HMI tags "PackTags"
   "PackTags.Admin.ProdProcessedCount[0].Count" : DInt = PLC PackTags.Admin.ProdProcessedCount[0].Count, 1 s   // Total Number of Products Through Machine / Número total de productos a través de la máquina
   "PackTags.Admin.ProdDefectiveCount[0].Count" : DInt = PLC PackTags.Admin.ProdDefectiveCount[0].Count, 1 s   // Total Number of Defective Products the Machine Processed (Reject Total ) / Número total de productos defectuosos procesados por la máquina (rechazo total)
   "PackTags.Admin.StopReason.ID" : DInt = PLC PackTags.Admin.StopReason.ID, 1 s   // Unique value assigned to each alarm
   "PackTags.Admin.StopReason.Value" : DInt = PLC PackTags.Admin.StopReason.Value, 1 s   // The Alarm Message number is a value that is associated to the alarm allowing for user specific detail or to break down the Alarm.ID to greater detail
   "PackTags.Admin.ProdProcessedCount[0].Unit" : String[5] = PLC PackTags.Admin.ProdProcessedCount[0].Unit, 1 s
   "PackTags.Admin.StatesDisabled" : DInt = PLC PackTags.Admin.StatesDisabled, 1 s
   "PackTags.Command.CmdChangeRequest" : Bool = PLC PackTags.Command.CmdChangeRequest, 1 s
   "PackTags.Command.CntrlCmd" : DInt = PLC PackTags.Command.CntrlCmd, 1 s
   "PackTags.Command.MachSpeed" : Real = PLC PackTags.Command.MachSpeed AT %DB1.DBD0, 1 s
   "PackTags.Command.UnitMode" : DInt = PLC PackTags.Command.UnitMode, 1 s
   "PackTags.Command.UnitModeChangeRequest" : Bool = PLC PackTags.Command.UnitModeChangeRequest, 1 s
   "PackML.remoteCommandEnable" : Bool = PLC PackML.remoteCommandEnable, 1 s
   "PackTags.Status.CurMachSpeed" : Real = PLC PackTags.Status.CurMachSpeed, 1 s
   "PackTags.Status.EquipmentInterlock.Blocked" : Bool = PLC PackTags.Status.EquipmentInterlock.Blocked, 1 s
   "PackTags.Status.EquipmentInterlock.Starved" : Bool = PLC PackTags.Status.EquipmentInterlock.Starved, 1 s
   "PackTags.Status.MachSpeed" : Real = PLC PackTags.Status.MachSpeed, 1 s
   "PackTags.Status.StateCurrent" : DInt = PLC PackTags.Status.StateCurrent, 500 ms
   "PackTags.Status.StateCurrentName" : String[16] = PLC PackTags.Status.StateCurrentName, 1 s
   "PackTags.Status.UnitModeCurrent" : DInt = PLC PackTags.Status.UnitModeCurrent, 1 s
   "PackTags.Status.UnitModeCurrentName" : String[18] = PLC PackTags.Status.UnitModeCurrentName, 1 s
   "PackML.Cmd.Mode.Maintenance" : Bool = PLC PackML.Cmd.Mode.Maintenance AT %DB1.DBX0.0, 1 s
   "PackML.Cmd.Mode.Manual" : Bool = PLC PackML.Cmd.Mode.Manual, 1 s
   "PackML.Cmd.Mode.Production" : Bool = PLC PackML.Cmd.Mode.Production, 1 s
   "PackML.Cmd.Mode.UserMode01" : Bool = PLC PackML.Cmd.Mode.UserMode01 AT %DB1.DBX0.0, 1 s
   "PackTags.Admin.AlarmExtent" : DInt = PLC PackTags.Admin.AlarmExtent, 1 s
   "PackTags.Admin.MachDesignSpeed" : Real = PLC PackTags.Admin.MachDesignSpeed AT %DB1.DBX0.0, 1 s
   "PackTags.Admin.ProdConsumedCount[0].AccCount" : DInt = PLC PackTags.Admin.ProdConsumedCount[0].AccCount, 1 s
   "PackTags.Admin.ProdConsumedCount[0].Count" : DInt = PLC PackTags.Admin.ProdConsumedCount[0].Count, 1 s
   "PackTags.Admin.ProdConsumedCount[0].Name" : String[24] = PLC PackTags.Admin.ProdConsumedCount[0].Name, 1 s
   "PackTags.Admin.ProdConsumedCount[0].Unit" : String[5] = PLC PackTags.Admin.ProdConsumedCount[0].Unit, 1 s
   "PackTags.Admin.ProdDefectiveCount[0].AccCount" : DInt = PLC PackTags.Admin.ProdDefectiveCount[0].AccCount, 1 s
   "PackTags.Admin.ProdDefectiveCount[0].Name" : String[24] = PLC PackTags.Admin.ProdDefectiveCount[0].Name, 1 s
   "PackTags.Admin.ProdDefectiveCount[0].Unit" : String[5] = PLC PackTags.Admin.ProdDefectiveCount[0].Unit, 1 s
   "PackTags.Admin.ProdProcessedCount[0].AccCount" : DInt = PLC PackTags.Admin.ProdProcessedCount[0].AccCount, 1 s
   "PackTags.Admin.ProdProcessedCount[0].Name" : String[24] = PLC PackTags.Admin.ProdProcessedCount[0].Name, 1 s
   "PackTags.Status.MaterialInterlock" : DWord = PLC PackTags.Status.MaterialInterlock AT %DB1.DBD0, 1 s

HMI tags "Tag table_PackTags_Times"
   "HMI_Data.resetPackMLTimers" : Bool = PLC HMI_Data.resetPackMLTimers, 500 ms   // Reset the PackML Timer values when set (1). / Restablezca los valores del temporizador PackML cuando se establece (1).
   "HMI_Data.modeCumulativeTime" : DInt = PLC HMI_Data.modeCumulativeTime, 1 s
   "HMI_Data.State_Current_Times[1]" : DInt = PLC HMI_Data.State_Current_Times[1], 1 s
   "HMI_Data.State_Current_Times[2]" : DInt = PLC HMI_Data.State_Current_Times[2], 1 s
   "HMI_Data.State_Current_Times[3]" : DInt = PLC HMI_Data.State_Current_Times[3], 1 s
   "HMI_Data.State_Current_Times[4]" : DInt = PLC HMI_Data.State_Current_Times[4], 1 s
   "HMI_Data.State_Current_Times[5]" : DInt = PLC HMI_Data.State_Current_Times[5], 1 s
   "HMI_Data.State_Current_Times[6]" : DInt = PLC HMI_Data.State_Current_Times[6], 1 s
   "HMI_Data.State_Current_Times[7]" : DInt = PLC HMI_Data.State_Current_Times[7], 1 s
   "HMI_Data.State_Current_Times[8]" : DInt = PLC HMI_Data.State_Current_Times[8], 1 s
   "HMI_Data.State_Current_Times[9]" : DInt = PLC HMI_Data.State_Current_Times[9], 1 s
   "HMI_Data.State_Current_Times[10]" : DInt = PLC HMI_Data.State_Current_Times[10], 1 s
   "HMI_Data.State_Current_Times[11]" : DInt = PLC HMI_Data.State_Current_Times[11], 1 s
   "HMI_Data.State_Current_Times[12]" : DInt = PLC HMI_Data.State_Current_Times[12], 1 s
   "HMI_Data.State_Current_Times[13]" : DInt = PLC HMI_Data.State_Current_Times[13], 1 s
   "HMI_Data.State_Current_Times[14]" : DInt = PLC HMI_Data.State_Current_Times[14], 1 s
   "HMI_Data.State_Current_Times[15]" : DInt = PLC HMI_Data.State_Current_Times[15], 1 s
   "HMI_Data.State_Current_Times[16]" : DInt = PLC HMI_Data.State_Current_Times[16], 1 s
   "HMI_Data.State_Current_Times[17]" : DInt = PLC HMI_Data.State_Current_Times[17], 1 s
   "HMI_Data.State_Cumulative_Times[1]" : DInt = PLC HMI_Data.State_Cumulative_Times[1], 1 s
   "HMI_Data.State_Cumulative_Times[2]" : DInt = PLC HMI_Data.State_Cumulative_Times[2], 1 s
   "HMI_Data.State_Cumulative_Times[3]" : DInt = PLC HMI_Data.State_Cumulative_Times[3], 1 s
   "HMI_Data.State_Cumulative_Times[4]" : DInt = PLC HMI_Data.State_Cumulative_Times[4], 1 s
   "HMI_Data.State_Cumulative_Times[5]" : DInt = PLC HMI_Data.State_Cumulative_Times[5], 1 s
   "HMI_Data.State_Cumulative_Times[6]" : DInt = PLC HMI_Data.State_Cumulative_Times[6], 1 s
   "HMI_Data.State_Cumulative_Times[7]" : DInt = PLC HMI_Data.State_Cumulative_Times[7], 1 s
   "HMI_Data.State_Cumulative_Times[8]" : DInt = PLC HMI_Data.State_Cumulative_Times[8], 1 s
   "HMI_Data.State_Cumulative_Times[9]" : DInt = PLC HMI_Data.State_Cumulative_Times[9], 1 s
   "HMI_Data.State_Cumulative_Times[10]" : DInt = PLC HMI_Data.State_Cumulative_Times[10], 1 s
   "HMI_Data.State_Cumulative_Times[11]" : DInt = PLC HMI_Data.State_Cumulative_Times[11], 1 s
   "HMI_Data.State_Cumulative_Times[12]" : DInt = PLC HMI_Data.State_Cumulative_Times[12], 1 s
   "HMI_Data.State_Cumulative_Times[13]" : DInt = PLC HMI_Data.State_Cumulative_Times[13], 1 s
   "HMI_Data.State_Cumulative_Times[14]" : DInt = PLC HMI_Data.State_Cumulative_Times[14], 1 s
   "HMI_Data.State_Cumulative_Times[15]" : DInt = PLC HMI_Data.State_Cumulative_Times[15], 1 s
   "HMI_Data.State_Cumulative_Times[16]" : DInt = PLC HMI_Data.State_Cumulative_Times[16], 1 s
   "HMI_Data.State_Cumulative_Times[17]" : DInt = PLC HMI_Data.State_Cumulative_Times[17], 1 s
   "PackTags.Admin.ModeCurrentTime[1]" : DInt = PLC PackTags.Admin.ModeCurrentTime[1], 1 s
   "PackTags.Admin.ModeCurrentTime[2]" : DInt = PLC PackTags.Admin.ModeCurrentTime[2], 1 s
   "PackTags.Admin.ModeCurrentTime[3]" : DInt = PLC PackTags.Admin.ModeCurrentTime[3], 1 s
   "PackTags.Admin.ModeCurrentTime[4]" : DInt = PLC PackTags.Admin.ModeCurrentTime[4], 1 s
   "PackTags.Admin.ModeCumulativeTime[1]" : DInt = PLC PackTags.Admin.ModeCumulativeTime[1], 1 s
   "PackTags.Admin.ModeCumulativeTime[2]" : DInt = PLC PackTags.Admin.ModeCumulativeTime[2], 1 s
   "PackTags.Admin.ModeCumulativeTime[3]" : DInt = PLC PackTags.Admin.ModeCumulativeTime[3], 1 s
   "PackTags.Admin.ModeCumulativeTime[4]" : DInt = PLC PackTags.Admin.ModeCumulativeTime[4], 1 s
   "PackTags.Admin.AccTimeSinceLastReset" : DInt = PLC PackTags.Admin.AccTimeSinceLastReset, 1 s

HMI tags "Tag table_Event_Warning_SortFilter"
   "HMI_Data.EMSortDisableWarning.EM00" : Bool = PLC HMI_Data.EMSortDisableWarning.EM00, 1 s   // If bool is reset, then EMxx sort filter is enabled, else it's disabled. / If bool is reset, then EMxx is sort filter is enabled, else it's disabled.
   "HMI_Data.EMSortDisableWarning.EM01" : Bool = PLC HMI_Data.EMSortDisableWarning.EM01, 1 s   // If bool is reset, then EMxx sort filter is enabled, else it's disabled. / If bool is reset, then EMxx is sort filter is enabled, else it's disabled.
   "HMI_Data.EMSortDisableWarning.EM02" : Bool = PLC HMI_Data.EMSortDisableWarning.EM02, 1 s   // If bool is reset, then EMxx sort filter is enabled, else it's disabled. / If bool is reset, then EMxx is sort filter is enabled, else it's disabled.
   "HMI_Data.EMSortDisableWarning.EM03" : Bool = PLC HMI_Data.EMSortDisableWarning.EM03, 1 s   // If bool is reset, then EMxx sort filter is enabled, else it's disabled. / If bool is reset, then EMxx is sort filter is enabled, else it's disabled.
   "HMI_Data.EMSortDisableWarning.EM04" : Bool = PLC HMI_Data.EMSortDisableWarning.EM04, 1 s   // If bool is reset, then EMxx sort filter is enabled, else it's disabled. / If bool is reset, then EMxx is sort filter is enabled, else it's disabled.
   "HMI_Data.EMSortDisableWarning.EM05" : Bool = PLC HMI_Data.EMSortDisableWarning.EM05, 1 s   // If bool is reset, then EMxx sort filter is enabled, else it's disabled. / If bool is reset, then EMxx is sort filter is enabled, else it's disabled.
   "HMI_Data.EMSortDisableWarning.EM06" : Bool = PLC HMI_Data.EMSortDisableWarning.EM06, 1 s   // If bool is reset, then EMxx sort filter is enabled, else it's disabled. / If bool is reset, then EMxx is sort filter is enabled, else it's disabled.
   "HMI_Data.EMSortDisableWarning.EM07" : Bool = PLC HMI_Data.EMSortDisableWarning.EM07, 1 s   // If bool is reset, then EMxx sort filter is enabled, else it's disabled. / If bool is reset, then EMxx is sort filter is enabled, else it's disabled.
   "HMI_Data.EMSortDisableWarning.EM08" : Bool = PLC HMI_Data.EMSortDisableWarning.EM08, 1 s   // If bool is reset, then EMxx sort filter is enabled, else it's disabled. / If bool is reset, then EMxx is sort filter is enabled, else it's disabled.
   "HMI_Data.EMSortDisableWarning.EM09" : Bool = PLC HMI_Data.EMSortDisableWarning.EM09, 1 s   // If bool is reset, then EMxx sort filter is enabled, else it's disabled. / If bool is reset, then EMxx is sort filter is enabled, else it's disabled.
   "HMI_Data.EMSortDisableWarning.EM10" : Bool = PLC HMI_Data.EMSortDisableWarning.EM10, 1 s   // If bool is reset, then EMxx sort filter is enabled, else it's disabled. / If bool is reset, then EMxx is sort filter is enabled, else it's disabled.
   "HMI_Data.EMSortDisableWarning.Unit" : Bool = PLC HMI_Data.EMSortDisableWarning.Unit, 1 s   // If bool is reset, then Unit sort filter is enabled, else it's disabled. / If bool is reset, then EMxx is sort filter is enabled, else it's disabled.

HMI tags "Tag table_Event_Warning"
   "HMI_Data.warningSortedList[0]" : CPG_typeEvent = PLC HMI_Data.warningSortedList[0], 1 s
   "HMI_Data.warningSortedList[1]" : CPG_typeEvent = PLC HMI_Data.warningSortedList[1], 1 s
   "HMI_Data.warningSortedList[2]" : CPG_typeEvent = PLC HMI_Data.warningSortedList[2], 1 s
   "HMI_Data.warningSortedList[3]" : CPG_typeEvent = PLC HMI_Data.warningSortedList[3], 1 s
   "HMI_Data.warningSortedList[4]" : CPG_typeEvent = PLC HMI_Data.warningSortedList[4], 1 s
   "HMI_Data.warningSortedList[5]" : CPG_typeEvent = PLC HMI_Data.warningSortedList[5], 1 s
   "HMI_Data.warningSortedList[6]" : CPG_typeEvent = PLC HMI_Data.warningSortedList[6], 1 s
   "HMI_Data.warningSortedList[7]" : CPG_typeEvent = PLC HMI_Data.warningSortedList[7], 1 s
   "HMI_Data.warningSortedList[8]" : CPG_typeEvent = PLC HMI_Data.warningSortedList[8], 1 s
   "HMI_Data.warningSortedList[9]" : CPG_typeEvent = PLC HMI_Data.warningSortedList[9], 1 s
   "HMI_Data.warningSortedList[10]" : CPG_typeEvent = PLC HMI_Data.warningSortedList[10], 1 s
   "HMI_Data.warningSortedList[11]" : CPG_typeEvent = PLC HMI_Data.warningSortedList[11], 1 s
   "HMI_Data.warningSortedList[12]" : CPG_typeEvent = PLC HMI_Data.warningSortedList[12], 1 s
   "HMI_Data.warningSortedList[13]" : CPG_typeEvent = PLC HMI_Data.warningSortedList[13], 1 s
   "HMI_Data.warningSortedList[14]" : CPG_typeEvent = PLC HMI_Data.warningSortedList[14], 1 s
   "HMI_Data.warningSortedList[15]" : CPG_typeEvent = PLC HMI_Data.warningSortedList[15], 1 s
   "HMI_Data.warningSortedList[16]" : CPG_typeEvent = PLC HMI_Data.warningSortedList[16], 1 s
   "HMI_Data.warningSortedList[17]" : CPG_typeEvent = PLC HMI_Data.warningSortedList[17], 1 s
   "HMI_Data.warningSortedList[18]" : CPG_typeEvent = PLC HMI_Data.warningSortedList[18], 1 s
   "HMI_Data.warningSortedList[19]" : CPG_typeEvent = PLC HMI_Data.warningSortedList[19], 1 s
   "HMI_Data.HMIWarningMsgScroll" : String[40] = PLC HMI_Data.HMIWarningMsgScroll, 1 s   // First Fault Messge - for HMI

HMI tags "Tag table_Event_Status"
   "Status.Summation.sts_Events[0]" : CPG_typeEvent = PLC Status.Summation.sts_Events[0], 1 s
   "Status.Summation.sts_Events[1]" : CPG_typeEvent = PLC Status.Summation.sts_Events[1], 1 s
   "Status.Summation.sts_Events[2]" : CPG_typeEvent = PLC Status.Summation.sts_Events[2], 1 s
   "Status.Summation.sts_Events[3]" : CPG_typeEvent = PLC Status.Summation.sts_Events[3], 1 s
   "Status.Summation.sts_Events[4]" : CPG_typeEvent = PLC Status.Summation.sts_Events[4], 1 s
   "Status.Summation.sts_Events[5]" : CPG_typeEvent = PLC Status.Summation.sts_Events[5], 1 s
   "Status.Summation.sts_Events[6]" : CPG_typeEvent = PLC Status.Summation.sts_Events[6], 1 s
   "Status.Summation.sts_Events[7]" : CPG_typeEvent = PLC Status.Summation.sts_Events[7], 1 s

HMI tags "Tag table_Event_AlarmHistory"
   "PackTags.Admin.AlarmHistory[0]" : CPG_typeEvent = PLC PackTags.Admin.AlarmHistory[0], 1 s
   "PackTags.Admin.AlarmHistory[1]" : CPG_typeEvent = PLC PackTags.Admin.AlarmHistory[1], 1 s
   "PackTags.Admin.AlarmHistory[2]" : CPG_typeEvent = PLC PackTags.Admin.AlarmHistory[2], 1 s
   "PackTags.Admin.AlarmHistory[3]" : CPG_typeEvent = PLC PackTags.Admin.AlarmHistory[3], 1 s
   "PackTags.Admin.AlarmHistory[4]" : CPG_typeEvent = PLC PackTags.Admin.AlarmHistory[4], 1 s
   "PackTags.Admin.AlarmHistory[5]" : CPG_typeEvent = PLC PackTags.Admin.AlarmHistory[5], 1 s
   "PackTags.Admin.AlarmHistory[6]" : CPG_typeEvent = PLC PackTags.Admin.AlarmHistory[6], 1 s
   "PackTags.Admin.AlarmHistory[7]" : CPG_typeEvent = PLC PackTags.Admin.AlarmHistory[7], 1 s
   "PackTags.Admin.AlarmHistory[8]" : CPG_typeEvent = PLC PackTags.Admin.AlarmHistory[8], 1 s
   "PackTags.Admin.AlarmHistory[9]" : CPG_typeEvent = PLC PackTags.Admin.AlarmHistory[9], 1 s

HMI tags "Tag table_Event_Alarm_SortFilter"
   "HMI_Data.EM_SortDisable_Alarm.Unit" : Bool = PLC HMI_Data.EM_SortDisable_Alarm.Unit, 1 s   // If bool is reset, then Unit sort filter is enabled, else it's disabled. / If bool is reset, then EMxx is sort filter is enabled, else it's disabled.
   "HMI_Data.EM_SortDisable_Alarm.EM10" : Bool = PLC HMI_Data.EM_SortDisable_Alarm.EM10, 1 s   // If bool is reset, then EMxx sort filter is enabled, else it's disabled. / If bool is reset, then EMxx is sort filter is enabled, else it's disabled.
   "HMI_Data.EM_SortDisable_Alarm.EM09" : Bool = PLC HMI_Data.EM_SortDisable_Alarm.EM09, 1 s   // If bool is reset, then EMxx sort filter is enabled, else it's disabled. / If bool is reset, then EMxx is sort filter is enabled, else it's disabled.
   "HMI_Data.EM_SortDisable_Alarm.EM08" : Bool = PLC HMI_Data.EM_SortDisable_Alarm.EM08, 1 s   // If bool is reset, then EMxx sort filter is enabled, else it's disabled. / If bool is reset, then EMxx is sort filter is enabled, else it's disabled.
   "HMI_Data.EM_SortDisable_Alarm.EM07" : Bool = PLC HMI_Data.EM_SortDisable_Alarm.EM07, 1 s   // If bool is reset, then EMxx sort filter is enabled, else it's disabled. / If bool is reset, then EMxx is sort filter is enabled, else it's disabled.
   "HMI_Data.EM_SortDisable_Alarm.EM06" : Bool = PLC HMI_Data.EM_SortDisable_Alarm.EM06, 1 s   // If bool is reset, then EMxx sort filter is enabled, else it's disabled. / If bool is reset, then EMxx is sort filter is enabled, else it's disabled.
   "HMI_Data.EM_SortDisable_Alarm.EM05" : Bool = PLC HMI_Data.EM_SortDisable_Alarm.EM05, 1 s   // If bool is reset, then EMxx sort filter is enabled, else it's disabled. / If bool is reset, then EMxx is sort filter is enabled, else it's disabled.
   "HMI_Data.EM_SortDisable_Alarm.EM04" : Bool = PLC HMI_Data.EM_SortDisable_Alarm.EM04, 1 s   // If bool is reset, then EMxx sort filter is enabled, else it's disabled. / If bool is reset, then EMxx is sort filter is enabled, else it's disabled.
   "HMI_Data.EM_SortDisable_Alarm.EM03" : Bool = PLC HMI_Data.EM_SortDisable_Alarm.EM03, 1 s   // If bool is reset, then EMxx sort filter is enabled, else it's disabled. / If bool is reset, then EMxx is sort filter is enabled, else it's disabled.
   "HMI_Data.EM_SortDisable_Alarm.EM02" : Bool = PLC HMI_Data.EM_SortDisable_Alarm.EM02, 1 s   // If bool is reset, then EMxx sort filter is enabled, else it's disabled. / If bool is reset, then EMxx is sort filter is enabled, else it's disabled.
   "HMI_Data.EM_SortDisable_Alarm.EM01" : Bool = PLC HMI_Data.EM_SortDisable_Alarm.EM01, 1 s   // If bool is reset, then EMxx sort filter is enabled, else it's disabled. / If bool is reset, then EMxx is sort filter is enabled, else it's disabled.
   "HMI_Data.EM_SortDisable_Alarm.EM00" : Bool = PLC HMI_Data.EM_SortDisable_Alarm.EM00, 1 s   // If bool is reset, then EMxx sort filter is enabled, else it's disabled. / If bool is reset, then EMxx is sort filter is enabled, else it's disabled.
   "HMI_Data.alarmFilter.cfgFilterCategory" : Int = PLC HMI_Data.alarmFilter.cfgFilterCategory, 1 s   // HMI - Alarm SortFilter - Filter Category #
   "HMI_Data.alarmFilter.cfgTimeSortDirection" : Bool = PLC HMI_Data.alarmFilter.cfgTimeSortDirection, 1 s   // HMI - Alarm SortFilter - Sort by Category
   "HMI_Data.alarmFilter.cmdFilterActiveEvents" : Bool = PLC HMI_Data.alarmFilter.cmdFilterActiveEvents, 1 s   // HMI - Alarm SortFilter - Filter Active Events
   "HMI_Data.alarmFilter.cmdFilterCategory" : Bool = PLC HMI_Data.alarmFilter.cmdFilterCategory, 1 s   // HMI - Alarm SortFilter - Filter Category
   "HMI_Data.alarmFilter.cmdSortCategory" : Bool = PLC HMI_Data.alarmFilter.cmdSortCategory, 1 s   // HMI - Alarm SortFilter - Sort by Time

HMI tags "Tag table_Event_Alarm"
   "PackTags.Admin.StopReason.Message" : String[60] = PLC PackTags.Admin.StopReason.Message, 1 s   // Message of alarm = prefix message + alarm message / Message OF alarm = prefix message + alarm message
   "HMI_Data.alarmSortedList[0]" : CPG_typeEvent = PLC HMI_Data.alarmSortedList[0], 1 s
   "HMI_Data.alarmSortedList[1]" : CPG_typeEvent = PLC HMI_Data.alarmSortedList[1], 1 s
   "HMI_Data.alarmSortedList[2]" : CPG_typeEvent = PLC HMI_Data.alarmSortedList[2], 1 s
   "HMI_Data.alarmSortedList[3]" : CPG_typeEvent = PLC HMI_Data.alarmSortedList[3], 1 s
   "HMI_Data.alarmSortedList[4]" : CPG_typeEvent = PLC HMI_Data.alarmSortedList[4], 1 s
   "HMI_Data.alarmSortedList[5]" : CPG_typeEvent = PLC HMI_Data.alarmSortedList[5], 1 s
   "HMI_Data.alarmSortedList[6]" : CPG_typeEvent = PLC HMI_Data.alarmSortedList[6], 1 s
   "HMI_Data.alarmSortedList[7]" : CPG_typeEvent = PLC HMI_Data.alarmSortedList[7], 1 s
   "HMI_Data.alarmSortedList[8]" : CPG_typeEvent = PLC HMI_Data.alarmSortedList[8], 1 s
   "HMI_Data.alarmSortedList[9]" : CPG_typeEvent = PLC HMI_Data.alarmSortedList[9], 1 s
   "HMI_Data.alarmSortedList[10]" : CPG_typeEvent = PLC HMI_Data.alarmSortedList[10], 1 s
   "HMI_Data.alarmSortedList[11]" : CPG_typeEvent = PLC HMI_Data.alarmSortedList[11], 1 s
   "HMI_Data.alarmSortedList[12]" : CPG_typeEvent = PLC HMI_Data.alarmSortedList[12], 1 s
   "HMI_Data.alarmSortedList[13]" : CPG_typeEvent = PLC HMI_Data.alarmSortedList[13], 1 s
   "HMI_Data.alarmSortedList[14]" : CPG_typeEvent = PLC HMI_Data.alarmSortedList[14], 1 s
   "HMI_Data.alarmSortedList[15]" : CPG_typeEvent = PLC HMI_Data.alarmSortedList[15], 1 s
   "HMI_Data.alarmSortedList[16]" : CPG_typeEvent = PLC HMI_Data.alarmSortedList[16], 1 s
   "HMI_Data.alarmSortedList[17]" : CPG_typeEvent = PLC HMI_Data.alarmSortedList[17], 1 s
   "HMI_Data.alarmSortedList[18]" : CPG_typeEvent = PLC HMI_Data.alarmSortedList[18], 1 s
   "HMI_Data.alarmSortedList[19]" : CPG_typeEvent = PLC HMI_Data.alarmSortedList[19], 1 s
   "PackTags.Admin.WarningExtent" : DInt = PLC PackTags.Admin.WarningExtent, 1 s

HMI tags "Tag table_EM_CM_Module Active"
   "EM00.PackML_Sts.Unit.moduleActive" : Bool = PLC EM00.PackML_Sts.Unit.moduleActive, 1 s   // Module Active Bit
   "EM01.PackML_Sts.Unit.moduleActive" : Bool = PLC EM01.PackML_Sts.Unit.moduleActive, 1 s   // Module Active Bit
   "UN.PackML_Sts.moduleActive" : Bool = PLC UN.PackML_Sts.moduleActive, 1 s   // Module Active Bit
   "EM02.PackML_Sts.Unit.moduleActive" : Bool = PLC EM02.PackML_Sts.Unit.moduleActive, 1 s

HMI tags "Tag table_HMI tags"
   "HMI_Data.ModeNames" : Array [0..4] of String[18] = PLC HMI_Data.ModeNames, 1 s
   "HMI_Data.StateNames" : Array [0..17] of String[16] = PLC HMI_Data.StateNames, 1 s
   "HMI_Data.languageSelected" : Int = PLC HMI_Data.languageSelected, 1 s   // This is the value of the language selected in the HMI (0=English, 1=DE, 2=SP, 3 / This is the value of the language selected in the HMI (0=English, 1=SP, 2=DE, 3
   "HMI_Data.CMDs.PB_Abort" : Bool = PLC HMI_Data.CMDs.PB_Abort, 1 s
   "HMI_Data.CMDs.PB_Complete" : Bool = PLC HMI_Data.CMDs.PB_Complete, 1 s
   "HMI_Data.CMDs.PB_Hold" : Bool = PLC HMI_Data.CMDs.PB_Hold, 1 s
   "HMI_Data.CMDs.PB_Reset" : Bool = PLC HMI_Data.CMDs.PB_Reset, 1 s
   "HMI_Data.CMDs.PB_Start" : Bool = PLC HMI_Data.CMDs.PB_Start, 1 s
   "HMI_Data.CMDs.PB_Stop" : Bool = PLC HMI_Data.CMDs.PB_Stop, 1 s
   "HMI_Data.CMDs.PB_EStop" : Bool = PLC HMI_Data.CMDs.PB_EStop, 1 s

HMI tags "Tag table_OEE_PWA"
   "PackML.OEE.realTime" : Real = PLC PackML.OEE.realTime, 1 s   // Real-Time OEE value / Echtzeit OEE Wert
   "PackML.OEE.availability" : Real = PLC PackML.OEE.availability, 1 s
   "PackML.OEE.performance" : Real = PLC PackML.OEE.performance, 1 s
   "PackML.OEE.quality" : Real = PLC PackML.OEE.quality, 1 s

HMI tags "Tag table_Recipes"
   "CPG_Recipe_Management.HMI_Command.Change.cancel" : Bool = PLC RecipeManagement.HMI_Command.Change.cancel, 1 s
   "CPG_Recipe_Management.HMI_Command.Change.changeCmd" : Bool = PLC RecipeManagement.HMI_Command.Change.changeCmd, 1 s
   "CPG_Recipe_Management.HMI_Command.Change.changeID" : Int = PLC RecipeManagement.HMI_Command.Change.changeID, 1 s
   "CPG_Recipe_Management.HMI_Command.Change.request" : Bool = PLC RecipeManagement.HMI_Command.Change.request, 1 s
   "CPG_Recipe_Management.HMI_Command.Delete.cancel" : Bool = PLC RecipeManagement.HMI_Command.Delete.cancel, 1 s
   "CPG_Recipe_Management.HMI_Command.Delete.deleteCmd" : Bool = PLC RecipeManagement.HMI_Command.Delete.deleteCmd, 1 s
   "CPG_Recipe_Management.HMI_Command.Delete.deleteID" : Int = PLC RecipeManagement.HMI_Command.Delete.deleteID, 1 s
   "CPG_Recipe_Management.HMI_Command.Delete.request" : Bool = PLC RecipeManagement.HMI_Command.Delete.request, 1 s
   "CPG_Recipe_Management.HMI_Command.Save.cancel" : Bool = PLC RecipeManagement.HMI_Command.Save.cancel, 1 s
   "CPG_Recipe_Management.HMI_Command.Save.request" : Bool = PLC RecipeManagement.HMI_Command.Save.request, 1 s
   "CPG_Recipe_Management.HMI_Command.Save.saveAsCmd" : Bool = PLC RecipeManagement.HMI_Command.Save.saveAsCmd, 1 s
   "CPG_Recipe_Management.HMI_Command.Save.saveAsDestinationID" : Int = PLC RecipeManagement.HMI_Command.Save.saveAsDestinationID, 1 s
   "CPG_Recipe_Management.HMI_Command.Save.saveAsNewName" : String[60] = PLC RecipeManagement.HMI_Command.Save.saveAsNewName, 1 s
   "CPG_Recipe_Management.HMI_Indicator.changeConfirm" : Bool = PLC RecipeManagement.HMI_Indicator.changeConfirm, 1 s
   "CPG_Recipe_Management.HMI_Indicator.deleteConfirm" : Bool = PLC RecipeManagement.HMI_Indicator.deleteConfirm, 1 s
   "CPG_Recipe_Management.HMI_Indicator.saveAsConfirm" : Bool = PLC RecipeManagement.HMI_Indicator.saveAsConfirm, 1 s
   "CPG_Recipe_Management.HMI_Command.Copy.cancel" : Bool = PLC RecipeManagement.HMI_Command.Copy.cancel, 1 s
   "CPG_Recipe_Management.HMI_Command.Copy.copyCmd" : Bool = PLC RecipeManagement.HMI_Command.Copy.copyCmd, 1 s
   "CPG_Recipe_Management.HMI_Command.Copy.copyDestinationID" : Int = PLC RecipeManagement.HMI_Command.Copy.copyDestinationID, 1 s
   "CPG_Recipe_Management.HMI_Command.Copy.copyNewName" : String[60] = PLC RecipeManagement.HMI_Command.Copy.copyNewName, 1 s
   "CPG_Recipe_Management.HMI_Command.Copy.copySourceID" : Int = PLC RecipeManagement.HMI_Command.Copy.copySourceID, 1 s
   "CPG_Recipe_Management.HMI_Command.Copy.request" : Bool = PLC RecipeManagement.HMI_Command.Copy.request, 1 s
   "CPG_Recipe_Management.HMI_Command.Save.saveCmd" : Bool = PLC RecipeManagement.HMI_Command.Save.saveCmd, 1 s
   "CPG_Recipe_Management.HMI_Indicator.copyConfirm" : Bool = PLC RecipeManagement.HMI_Indicator.copyConfirm, 1 s
   "CPG_RecipeCfg.recipeControl" : CPG_typeRecipeControl = PLC RecipeCfg.recipeControl, 1 s
   "CPG_Recipe_Management.HMI_Indicator.changeErr" : Bool = PLC RecipeManagement.HMI_Indicator.changeErr AT %DB1.DBW0, 1 s
   "CPG_Recipe_Management.HMI_Indicator.saveAsErr" : Bool = PLC RecipeManagement.HMI_Indicator.saveAsErr AT %DB1.DBX0.0, 1 s
   "CPG_Recipe_Management.HMI_Indicator.copyErr" : Bool = PLC RecipeManagement.HMI_Indicator.copyErr AT %DB1.DBX0.0, 1 s
   "CPG_Recipe_Management.HMI_Indicator.deleteErr" : Bool = PLC RecipeManagement.HMI_Indicator.deleteErr AT %DB1.DBX0.0, 1 s
   "CPG_Recipe_Management.recipeArrayTimes" : Array [0..19] of Time = PLC RecipeManagement.recipeArrayTimes AT %DB1.DBW0, 1 s
   "CPG_Recipe_Management.recipeArraySaves" : Array [0..19] of DTL = PLC RecipeManagement.recipeArraySaves AT %DB1.DBX0.0, 1 s
   "CPG_Recipe_Management.recipeArrayNames" : Array [0..19] of String[60] = PLC RecipeManagement.recipeArrayNames AT %DB1.DBX0.0, 1 s
   "CPG_Recipe_Management.HMI_Command.resetAllTimes" : Bool = PLC RecipeManagement.HMI_Command.resetAllTimes, 1 s
   "CPG_Recipe_Management.setpointsArray_REAL[0]" : CPG_typeRecipeSetpoint_REAL = PLC RecipeManagement.setpointsArray_REAL[0] AT %DB1.DBX0.0, 1 s
   "CPG_Recipe_Management.setpointsArray_REAL[1]" : CPG_typeRecipeSetpoint_REAL = PLC RecipeManagement.setpointsArray_REAL[1] AT %DB1.DBX0.0, 1 s
   "CPG_Recipe_Management.setpointsArray_REAL[2]" : CPG_typeRecipeSetpoint_REAL = PLC RecipeManagement.setpointsArray_REAL[2] AT %DB1.DBX0.0, 1 s
   "CPG_Recipe_Management.setpointsArray_REAL[3]" : CPG_typeRecipeSetpoint_REAL = PLC RecipeManagement.setpointsArray_REAL[3] AT %DB1.DBX0.0, 1 s
   "CPG_Recipe_Management.setpointsArray_REAL[4]" : CPG_typeRecipeSetpoint_REAL = PLC RecipeManagement.setpointsArray_REAL[4] AT %DB1.DBX0.0, 1 s
   "CPG_Recipe_Management.setpointsArray_REAL[5]" : CPG_typeRecipeSetpoint_REAL = PLC RecipeManagement.setpointsArray_REAL[5] AT %DB1.DBX0.0, 1 s
   "CPG_Recipe_Management.setpointsArray_REAL[6]" : CPG_typeRecipeSetpoint_REAL = PLC RecipeManagement.setpointsArray_REAL[6] AT %DB1.DBX0.0, 1 s
   "CPG_Recipe_Management.setpointsArray_REAL[7]" : CPG_typeRecipeSetpoint_REAL = PLC RecipeManagement.setpointsArray_REAL[7] AT %DB1.DBX0.0, 1 s
   "CPG_Recipe_Management.setpointsArray_REAL[8]" : CPG_typeRecipeSetpoint_REAL = PLC RecipeManagement.setpointsArray_REAL[8] AT %DB1.DBX0.0, 1 s
   "CPG_Recipe_Management.setpointsArray_REAL[9]" : CPG_typeRecipeSetpoint_REAL = PLC RecipeManagement.setpointsArray_REAL[9] AT %DB1.DBX0.0, 1 s
   "CPG_Recipe_Management.setpointsArray_REAL[10]" : CPG_typeRecipeSetpoint_REAL = PLC RecipeManagement.setpointsArray_REAL[10] AT %DB1.DBX0.0, 1 s
   "CPG_Recipe_Management.setpointsArray_REAL[11]" : CPG_typeRecipeSetpoint_REAL = PLC RecipeManagement.setpointsArray_REAL[11] AT %DB1.DBX0.0, 1 s
   "CPG_Recipe_Management.setpointsArray_DINT[0]" : CPG_typeRecipeSetpoint_DINT = PLC RecipeManagement.setpointsArray_DINT[0], 1 s
   "CPG_Recipe_Management.setpointsArray_DINT[1]" : CPG_typeRecipeSetpoint_DINT = PLC RecipeManagement.setpointsArray_DINT[1], 1 s
   "CPG_Recipe_Management.setpointsArray_DINT[2]" : CPG_typeRecipeSetpoint_DINT = PLC RecipeManagement.setpointsArray_DINT[2], 1 s
   "CPG_Recipe_Management.setpointsArray_DINT[3]" : CPG_typeRecipeSetpoint_DINT = PLC RecipeManagement.setpointsArray_DINT[3], 1 s
   "CPG_Recipe_Management.setpointsArray_DINT[4]" : CPG_typeRecipeSetpoint_DINT = PLC RecipeManagement.setpointsArray_DINT[4], 1 s
   "CPG_Recipe_Management.setpointsArray_DINT[5]" : CPG_typeRecipeSetpoint_DINT = PLC RecipeManagement.setpointsArray_DINT[5], 1 s
   "CPG_Recipe_Management.setpointsArray_DINT[6]" : CPG_typeRecipeSetpoint_DINT = PLC RecipeManagement.setpointsArray_DINT[6], 1 s
   "CPG_Recipe_Management.setpointsArray_DINT[7]" : CPG_typeRecipeSetpoint_DINT = PLC RecipeManagement.setpointsArray_DINT[7], 1 s
   "CPG_Recipe_Management.setpointsArray_DINT[8]" : CPG_typeRecipeSetpoint_DINT = PLC RecipeManagement.setpointsArray_DINT[8], 1 s
   "CPG_Recipe_Management.setpointsArray_DINT[9]" : CPG_typeRecipeSetpoint_DINT = PLC RecipeManagement.setpointsArray_DINT[9], 1 s
   "CPG_Recipe_Management.setpointsArray_DINT[10]" : CPG_typeRecipeSetpoint_DINT = PLC RecipeManagement.setpointsArray_DINT[10], 1 s
   "CPG_Recipe_Management.setpointsArray_DINT[11]" : CPG_typeRecipeSetpoint_DINT = PLC RecipeManagement.setpointsArray_DINT[11], 1 s
   "CPG_Recipe_Management.setpointsArray_BOOL[0]" : CPG_typeRecipeSetpoint_BOOL = PLC RecipeManagement.setpointsArray_BOOL[0], 1 s
   "CPG_Recipe_Management.setpointsArray_BOOL[1]" : CPG_typeRecipeSetpoint_BOOL = PLC RecipeManagement.setpointsArray_BOOL[1], 1 s
   "CPG_Recipe_Management.setpointsArray_BOOL[2]" : CPG_typeRecipeSetpoint_BOOL = PLC RecipeManagement.setpointsArray_BOOL[2], 1 s
   "CPG_Recipe_Management.setpointsArray_BOOL[3]" : CPG_typeRecipeSetpoint_BOOL = PLC RecipeManagement.setpointsArray_BOOL[3], 1 s
   "CPG_Recipe_Management.setpointsArray_BOOL[4]" : CPG_typeRecipeSetpoint_BOOL = PLC RecipeManagement.setpointsArray_BOOL[4], 1 s
   "CPG_Recipe_Management.setpointsArray_BOOL[5]" : CPG_typeRecipeSetpoint_BOOL = PLC RecipeManagement.setpointsArray_BOOL[5], 1 s
   "CPG_Recipe_Management.setpointsArray_BOOL[6]" : CPG_typeRecipeSetpoint_BOOL = PLC RecipeManagement.setpointsArray_BOOL[6], 1 s
   "CPG_Recipe_Management.setpointsArray_BOOL[7]" : CPG_typeRecipeSetpoint_BOOL = PLC RecipeManagement.setpointsArray_BOOL[7], 1 s
   "CPG_Recipe_Management.setpointsArray_BOOL[8]" : CPG_typeRecipeSetpoint_BOOL = PLC RecipeManagement.setpointsArray_BOOL[8], 1 s
   "CPG_Recipe_Management.setpointsArray_BOOL[9]" : CPG_typeRecipeSetpoint_BOOL = PLC RecipeManagement.setpointsArray_BOOL[9], 1 s
   "CPG_Recipe_Management.setpointsArray_BOOL[10]" : CPG_typeRecipeSetpoint_BOOL = PLC RecipeManagement.setpointsArray_BOOL[10], 1 s
   "CPG_Recipe_Management.setpointsArray_BOOL[11]" : CPG_typeRecipeSetpoint_BOOL = PLC RecipeManagement.setpointsArray_BOOL[11], 1 s
   "CPG_Recipe_Management.setpointsArray_STRING[0]" : CPG_typeRecipeSetpoint_STRING = PLC RecipeManagement.setpointsArray_STRING[0] AT %DB1.DBW0, 1 s
   "CPG_Recipe_Management.setpointsArray_STRING[1]" : CPG_typeRecipeSetpoint_STRING = PLC RecipeManagement.setpointsArray_STRING[1] AT %DB1.DBW0, 1 s
   "CPG_Recipe_Management.setpointsArray_STRING[2]" : CPG_typeRecipeSetpoint_STRING = PLC RecipeManagement.setpointsArray_STRING[2] AT %DB1.DBW0, 1 s
   "CPG_Recipe_Management.setpointsArray_STRING[3]" : CPG_typeRecipeSetpoint_STRING = PLC RecipeManagement.setpointsArray_STRING[3] AT %DB1.DBW0, 1 s
   "CPG_Recipe_Management.setpointsArray_STRING[4]" : CPG_typeRecipeSetpoint_STRING = PLC RecipeManagement.setpointsArray_STRING[4] AT %DB1.DBW0, 1 s
   "CPG_Recipe_Management.setpointsArray_STRING[5]" : CPG_typeRecipeSetpoint_STRING = PLC RecipeManagement.setpointsArray_STRING[5] AT %DB1.DBW0, 1 s
   "CPG_Recipe_Management.setpointsArray_STRING[6]" : CPG_typeRecipeSetpoint_STRING = PLC RecipeManagement.setpointsArray_STRING[6] AT %DB1.DBW0, 1 s
   "CPG_Recipe_Management.setpointsArray_STRING[7]" : CPG_typeRecipeSetpoint_STRING = PLC RecipeManagement.setpointsArray_STRING[7] AT %DB1.DBW0, 1 s
   "CPG_Recipe_Management.setpointsArray_STRING[8]" : CPG_typeRecipeSetpoint_STRING = PLC RecipeManagement.setpointsArray_STRING[8] AT %DB1.DBW0, 1 s
   "CPG_Recipe_Management.setpointsArray_STRING[9]" : CPG_typeRecipeSetpoint_STRING = PLC RecipeManagement.setpointsArray_STRING[9] AT %DB1.DBW0, 1 s
   "CPG_Recipe_Management.setpointsArray_STRING[10]" : CPG_typeRecipeSetpoint_STRING = PLC RecipeManagement.setpointsArray_STRING[10] AT %DB1.DBW0, 1 s
   "CPG_Recipe_Management.setpointsArray_STRING[11]" : CPG_typeRecipeSetpoint_STRING = PLC RecipeManagement.setpointsArray_STRING[11] AT %DB1.DBW0, 1 s
   "CPG_Recipe_Management.setpointPopup_REAL" : CPG_typeRecipeSetpoint_REAL = PLC RecipeManagement.setpointPopup_REAL AT %DB1.DBW0, 1 s
   "CPG_Recipe_Management.setpointPopup_DINT" : CPG_typeRecipeSetpoint_DINT = PLC RecipeManagement.setpointPopup_DINT AT %DB1.DBW0, 1 s
   "CPG_Recipe_Management.setpointPopup_BOOL" : CPG_typeRecipeSetpoint_BOOL = PLC RecipeManagement.setpointPopup_BOOL, 1 s
   "CPG_Recipe_Management.setpointPopup_STRING" : CPG_typeRecipeSetpoint_STRING = PLC RecipeManagement.setpointPopup_STRING, 1 s
   "CPG_Recipe_Management.popupTrackers[0]" : Int = PLC RecipeManagement.popupTrackers[0], 1 s
   "CPG_Recipe_Management.popupTrackers[1]" : Int = PLC RecipeManagement.popupTrackers[1] AT %DB1.DBW0, 1 s
   "CPG_Recipe_Management.popupTrackers[2]" : Int = PLC RecipeManagement.popupTrackers[2] AT %DB1.DBW0, 1 s
   "CPG_Recipe_Management.popupTrackers[3]" : Int = PLC RecipeManagement.popupTrackers[3] AT %DB1.DBW0, 1 s
   "CPG_Recipe_Management.currentPages[0]" : Int = PLC RecipeManagement.currentPages[0] AT %DB1.DBW0, 1 s
   "CPG_Recipe_Management.currentPages[1]" : Int = PLC RecipeManagement.currentPages[1] AT %DB1.DBW0, 1 s
   "CPG_Recipe_Management.currentPages[2]" : Int = PLC RecipeManagement.currentPages[2] AT %DB1.DBW0, 1 s
   "CPG_Recipe_Management.currentPages[3]" : Int = PLC RecipeManagement.currentPages[3] AT %DB1.DBW0, 1 s
   "CPG_Recipe_Management.maxPages[0]" : Int = PLC RecipeManagement.maxPages[0] AT %DB1.DBW0, 1 s
   "CPG_Recipe_Management.maxPages[1]" : Int = PLC RecipeManagement.maxPages[1] AT %DB1.DBW0, 1 s
   "CPG_Recipe_Management.maxPages[2]" : Int = PLC RecipeManagement.maxPages[2] AT %DB1.DBW0, 1 s
   "CPG_Recipe_Management.maxPages[3]" : Int = PLC RecipeManagement.maxPages[3] AT %DB1.DBW0, 1 s
   "CPG_Recipe_Management.displayDisable_REAL" : Array [0..11] of Bool = PLC RecipeManagement.displayDisable_REAL AT %DB1.DBX0.0, 1 s
   "CPG_Recipe_Management.displayDisable_DINT" : Array [0..11] of Bool = PLC RecipeManagement.displayDisable_DINT AT %DB1.DBX0.0, 1 s
   "CPG_Recipe_Management.displayDisable_BOOL" : Array [0..11] of Bool = PLC RecipeManagement.displayDisable_BOOL AT %DB1.DBX0.0, 1 s
   "CPG_Recipe_Management.displayDisable_STRING" : Array [0..11] of Bool = PLC RecipeManagement.displayDisable_STRING, 1 s
   "CPG_Recipe_Management.currentPages[4]" : Int = PLC RecipeManagement.currentPages[4] AT %DB1.DBX0.0, 1 s
   "CPG_Recipe_Management.maxPages[4]" : Int = PLC RecipeManagement.maxPages[4] AT %DB1.DBW0, 1 s
   "CPG_Recipe_Management.recipeArrayNums" : Array [0..19] of Int = PLC RecipeManagement.recipeArrayNums AT %DB1.DBX0.0, 1 s
   "CPG_Recipe_Management.recipeArrayHide" : Array [0..19] of Bool = PLC RecipeManagement.recipeArrayHide AT %DB1.DBX0.0, 1 s

HMI tags "Pareto_Tags"
   "ParetoData_Reset" : Bool = PLC ParetoData.Reset, 1 s
   "ParetoData_totalStops" : Int = PLC ParetoData.totalStops AT %DB1.DBX0.0, 1 s
   "ParetoData_Sort" : Int = PLC ParetoData.Sort AT %DB1.DBW0, 1 s
   "ParetoData_totalUptime" : Real = PLC ParetoData.totalUptime AT %DB1.DBW0, 1 s
   "ParetoData_totalDowntime" : Real = PLC ParetoData.totalDowntime AT %DB1.DBD0, 1 s
   "ParetoData_totalTimeSinceReset" : Real = PLC ParetoData.totalTimeSinceReset AT %DB1.DBD0, 1 s
   "ParetoData_percentUptime" : Real = PLC ParetoData.percentUptime AT %DB1.DBD0, 1 s
   "ParetoData_MTTR" : Real = PLC ParetoData.MTTR AT %DB1.DBD0, 1 s
   "ParetoData_MTBF" : Real = PLC ParetoData.MTBF AT %DB1.DBD0, 1 s
   "ParetoData_alarmOccurrence[1]" : CPG_typePareto = PLC ParetoData.alarmOccurrence[1] AT %DB1.DBD0, 1 s
   "ParetoData_alarmOccurrence[2]" : CPG_typePareto = PLC ParetoData.alarmOccurrence[2] AT %DB1.DBD0, 1 s
   "ParetoData_alarmOccurrence[3]" : CPG_typePareto = PLC ParetoData.alarmOccurrence[3] AT %DB1.DBD0, 1 s
   "ParetoData_alarmOccurrence[4]" : CPG_typePareto = PLC ParetoData.alarmOccurrence[4] AT %DB1.DBD0, 1 s
   "ParetoData_alarmOccurrence[5]" : CPG_typePareto = PLC ParetoData.alarmOccurrence[5] AT %DB1.DBD0, 1 s
   "ParetoData_alarmOccurrence[6]" : CPG_typePareto = PLC ParetoData.alarmOccurrence[6] AT %DB1.DBD0, 1 s
   "ParetoData_alarmOccurrence[7]" : CPG_typePareto = PLC ParetoData.alarmOccurrence[7] AT %DB1.DBD0, 1 s
   "ParetoData_alarmOccurrence[8]" : CPG_typePareto = PLC ParetoData.alarmOccurrence[8] AT %DB1.DBD0, 1 s
   "ParetoData_alarmOccurrence[9]" : CPG_typePareto = PLC ParetoData.alarmOccurrence[9] AT %DB1.DBD0, 1 s
   "ParetoData_alarmOccurrence[10]" : CPG_typePareto = PLC ParetoData.alarmOccurrence[10] AT %DB1.DBD0, 1 s

HMI tags "Tag table_Labeler"
   "HMI_Data_Custom.MachineSpeed_SP" : Real = PLC HMI_Data_Custom.machineSpeedSP, 1 s
   "HMI_Data_Custom.MachineSpeed_PV" : Real = PLC HMI_Data_Custom.machineSpeedPV, 1 s
   "HMI_Data_CPG.CMDs.PB_EStop" : Bool = PLC HMI_Data.CMDs.PB_EStop, 1 s

HMI tags "Constants"
   "bo_TRUE" : Bool, internal
   "bo_FALSE" : Bool, internal
   "i16_1000_MachineControl_SecondNavMaxTopics" : Int, internal
   "i16_2000_Settings_SecondNavMaxTopics" : Int, internal
   "i16_3000_Alarms&Events_SecondNavMaxTopics" : Int, internal
   "i16_4000_Statistics_SecondNavMaxTopics" : Int, internal
   "i16_5000_Manual_SecondNavMaxTopics" : Int, internal
   "i16_6000_Diagnostics_SecondNavMaxTopics" : Int, internal
   "i16_7000_Formats_SecondNavMaxTopics" : Int, internal

HMI tags "Systemfunction"
   "i16_Settings_CurDisplayBrightness" : Int, internal
   "HMI_Data.HMICurrentScreenID" : Int = PLC HMI_Data.HMICurrentScreenID AT %MW0, 1 s   // Internal tag, but has to be connected to a PLC
   "str_System_CurUser" : WString[20], internal
   "bo_System_BaseScreenLocked" : Bool, internal
   "str_Diagnostic_WebURL" : WString[255], internal
   "i16_Format_CurSelectedRecipeID" : Int, internal
   "i16_Format_CurSelectedRecSetID" : Int, internal
   "bo_System_PLCConnectionOK" : Bool, internal
   "arr_System_PrevScreenStorage" : Array [0..10] of Int, internal
   "bo_System_PrevScreenActive" : Bool, internal
   "i16_System_PrevScreenPointer" : Int, internal
   "dat_Settings_NewDateTime" : DateTime, internal
   "i16_Format_RecipeTag" : Int, internal
   "i16_PLCConnectionOK" : Int, internal

text list "LPMLV30_States": 0 'Undefined / Indefinido'; 1 'Clearing'; 2 'Stopped / Detenerped'; 3 'Starting / Comienzoing'; 4 'Idle / Ocioso'; 5 'Suspended'; 6 'Execute'; 7 'Stopping / Detenerping'; 8 'Aborting / Abortaring'; 9 'Aborted / Abortared'; 10 'Holding'; 11 'Held / Retenida'; 12 'Unholding / Desactivar'; 13 'Suspending'; 14 'Unsuspending'; 15 'Resetting / Restablecer'; 16 'Completing'; 17 'Complete'; 0 'Undefined'

text list "LPMLV30_CntrlCmd": 1 'Reset / Reiniciar'; 2 'Start / Comienzo'; 3 'Stop / Detener'; 4 'Hold'; 5 'Unhold'; 6 'Suspend'; 7 'Unsuspend'; 8 'Abort / Abortar'; 9 'Clear'; 0 'Undefined / Indefinido'; 10 'Complete'; 0 'Undefined'

text list "LPMLV30_Message": 0 '16#xx: unknown status value'; 1 '16#01: unitMode changed successfully'; 2 '16#02: state changed successfully'; 128 '16#80: unitMode invalid'; 129 '16#81: cntrlCmd undefined'; 130 '16#82: requested unitMode not configured'; 131 '16#83: unitMode transition not allowed'; 132 '16#84: cntrlCmd in this state not allowed'; 133 '16#85: SC in this state not allowed'; 134 '16#86: state configuration was forced to OMAC standard'; 135 '16#87: wrong use of boolean interface'; 0 '16#00: - - -'

text list "LPMLV30_UnitModes": 0..1 'Invalid / Indefinido'; 1 'Production / Produktion / Produccion'; 2 'Maintenance / Wartung / Mantenimiento'; 3 'Manual / Hand / Manual (Factory)'; 4 'User Mode 1 / Benutzermode 1 / Change over'; 0 'Invalid'; 5 'User Mode 2'; 6 'User Mode 3'; 7 'User Mode 4'; 8 'User Mode 5'; 9 'User Mode 6'; 10 'User Mode 7'; 11 'User Mode 8'; 12 'User Mode 9'; 13 'User Mode 10'; 14 'User Mode 11'; 15 'User Mode 12'; 16 'User Mode 13'; 17 'User Mode 14'; 18 'User Mode 15'; 19 'User Mode 16'; 20 'User Mode 17'; 21 'User Mode 18'; 22 'User Mode 19'; 23 'User Mode 20'; 24 'User Mode 21'; 25 'User Mode 22'; 26 'User Mode 23'; 27 'User Mode 24'; 28 'User Mode 25'; 29 'User Mode 26'; 30 'User Mode 27'; 31 'User Mode 28'

text list "ScreenName": 0 'Runtime Start... / Runtime Comienzo...'; 1001 'Overview / Übersicht / Equipment View 1'; 1041 'Up & Downstream'; 1081 'OMAC State Model / OMAC Statusmodell'; 2041 'System Functions / Systemfunktionen / Funciones del sistema'; 2081 'User Management / Benutzerverwaltung / User Managment'; 3001 'Event Overview / Ereignisübersicht / TR88 Resumen del evento'; 3041 'Alarm Events / Alarmmeldungen / TR88 Alarmas activas'; 3081 'Warning Events / Warnmeldungen / Advertencias activas TR88'; 3121 'HMI Events / HMI Meldungen / HMI Messages'; 6001 'System Diagnostic / Systemdiagnose / Diagnostico del sistema'; 6041 'Web Diagnostic / Webdiagnose / Diagnóstico web'; 7001 'Format Management / Rezepturverwaltung'; 1121 'OMAC PackTags / PackTags'; 1161 'OMAC Times / OMAC Zeiten / Times / OEE'; 1241 'Manual Commands / Manuelle Kommandos / Topic6'; 1201 'OEE'; -1 '?????'; 2001 'Einstellungen / Settings'; 3161 'Pareto Alarmdaten / Pareto Alarm Data'; 7041 'REAL Sollwerte / Recipe Setpoints REAL'; 7081 'DINT Sollwerte / Recipe Setpoints DINT'; 7121 'BOOL Sollwerte / Recipe Setpoints BOOL'; 7161 'STRING Sollwerte / Recipe Setpoints STRING'

text list "CPG_CategoryList": 0 '(0) - E-Stop / (0) - Molestar'; 1 '(1) - Abort / (1) - Abortar'; 2 '(2) - Stop / (2) - Detener'; 3 '(3) - Stop / (3) - Detener'; 4 '(4) - Stop / (4) - Detener'; 5 '(5) -'; 6 '(6) -'; 7 '(7) - Held / (7) - Retenida'; 8 '(8) - Blocked / (8) - Obstruido'; 9 '(9) - Starved / (9) - Famélico'

text list "MaterialInterlock_LabelSupply_Ready": 0 'Not Ready / No esta listo / Nicht bereit'; 1 'Ready / Listo / Bereit'

text list "MaterialInterlock_LabelSupply_NotLow": 0 'Low / Bajo / Niedrig'; 1 'Not Low / No bajo / Nicht niedrig'

text list "Local_Remote_Control": 0 'Local Control Only Control local Solamente Lokale Kontrolle freigegegeben'; 1 'Remote Control Enabled Control remoto Habilitado Remote Control freigegeben'

text list "MaterialInterlock_BottleSupply_NotLow": 0 'Low / Bajo / Niedrig'; 1 'Not Low / No bajo / Nicht niedrig'

text list "MaterialInterlock_BottleSupply_Ready": 0 'Not Ready / No esta listo / Nicht bereit'; 1 'Ready / Listo / Bereit'

text list "Pareto_Sort": 0 'Gesamt-Unproduktiv / Total Downtime'; 1 'Anteil % / Percentage Occurred'; 2 'Anzahl / Times Occurred'; 3 'MTTR'

graphic list "PLCConnectionStatus": 0 'icn-status-notOK-32x32'; 1 'icn-status-OK-32x32'

graphic list "MaterialInterlocksReadyOrNotLow": 0 'PilotLight_Square_R_On_256c'; 1 'PilotLight_Square_GN_On_256c'

recipe "Recipe": Recipe_element_1 <- "i16_Format_RecipeTag"

screen "Startup Screen" 1280x715, template "1xxx_MachineControl"
   on GenerateScreen: "sub_RuntimeStart"()
   TextField "txtInfo" at 5,5 size 1095x615; Text 'The runtime is starting. Please wait... / Die Runtime wird gestartet. Bitte warten...'

screen "1001_EquipmentView1" 1280x715, template "1xxx_MachineControl"
   TextField "fraOperatorInformation" at 15,446 size 788x164; Text 'Operator Information / Bedienerinformationen / Información del operador:'
   TextField "txtActiveEventsID" at 50,475 size 55x25; Text 'ID / ID:'
   TextField "txtActiveEventsMessage" at 105,475 size 490x25; Text 'Message / Meldung / Mensaje:'
   TextField "txtActiveEventsTimeIn" at 595,475 size 200x25; Text 'Time In / Gekommen / Tiempo en:'
   TextField "txtActiveEventsRow1" at 25,500 size 25x25; Text '1'
   TextField "txtActiveEventsRow2" at 25,525 size 25x25; Text '2'
   TextField "txtActiveEventsRow3" at 25,550 size 25x25; Text '3'
   TextField "txtActiveEventsRow4" at 25,575 size 25x25; Text '4'
   ScreenModuleView "fcpActiveEventsRow1-2" at 50,500 size 745x51; ScreenModuleType ""
      Guid_{11997190-459382} <- "Status.Summation.sts_Events[0]"
      Guid_{11997190-459405} <- "Status.Summation.sts_Events[1]"
   ScreenModuleView "fcpActiveEventsRow3-4" at 50,550 size 745x51; ScreenModuleType ""
      Guid_{11997190-459382} <- "Status.Summation.sts_Events[2]"
      Guid_{11997190-459405} <- "Status.Summation.sts_Events[3]"
   Rectangle "recBaseScreenLocked" at 0,0 size 1280x708
      Visibility <- "bo_System_BaseScreenLocked"

screen "1041_Up&Downstream" 1280x715, template "1xxx_MachineControl"
   Rectangle "recBaseScreenLocked" at 0,0 size 1280x708
      Visibility <- "bo_System_BaseScreenLocked"
   TextField "fraMaterielSupply" at 15,15 size 536x173; Text 'Material Supply / Materialversorgung / Suministro de material:'
   TextField "txtMaterialSupply2" at 25,120 size 220x25; Text 'Material Supply #2: / Materialversorgung #2: / Materia prima # 1 vacía .....'
   TextField "txtMaterialSupply1" at 25,55 size 220x25; Text 'Material Supply #1: / Materialversorgung #1: / Materia prima # 1 vacía .....'
   GraphicIOField "valOutput1MaterialSupply1Ready" at 250,55 size 25x25; PictureOn "PilotLight_Square_GN_On_256c"; PictureOff "PilotLight_Square_R_On_256c"; PictureList "MaterialInterlocksReadyOrNotLow"
      ProcessValue <- "PackTags.Status.MaterialInterlock"
   GraphicIOField "valOutput1MaterialSupply1Low" at 250,86 size 25x25; PictureOn "PilotLight_Square_GN_On_256c"; PictureOff "PilotLight_Square_R_On_256c"; PictureList "MaterialInterlocksReadyOrNotLow"
      ProcessValue <- "PackTags.Status.MaterialInterlock"
   SymbolicIOField "valOutput2MaterialSupply1Ready" at 278,55 size 220x25; TextOn '1'; TextOff '0'; TextList "MaterialInterlock_BottleSupply_Ready"
      ProcessValue <- "PackTags.Status.MaterialInterlock"
   SymbolicIOField "valOutput2MaterialSupply1Low" at 279,85 size 220x25; TextOn '1'; TextOff '0'; TextList "MaterialInterlock_BottleSupply_NotLow"
      ProcessValue <- "PackTags.Status.MaterialInterlock"
   GraphicIOField "valOutput1MaterialSupply2Ready" at 250,120 size 25x25; PictureOn "PilotLight_Square_GN_On_256c"; PictureOff "PilotLight_Square_R_On_256c"; PictureList "MaterialInterlocksReadyOrNotLow"
      ProcessValue <- "PackTags.Status.MaterialInterlock"
   GraphicIOField "valOutput1MaterialSupply2Low" at 250,151 size 25x25; PictureOn "PilotLight_Square_GN_On_256c"; PictureOff "PilotLight_Square_R_On_256c"; PictureList "MaterialInterlocksReadyOrNotLow"
      ProcessValue <- "PackTags.Status.MaterialInterlock"
   SymbolicIOField "valOutput2MaterialSupply2Ready" at 279,120 size 220x25; TextOn '1'; TextOff '0'; TextList "MaterialInterlock_LabelSupply_Ready"
      ProcessValue <- "PackTags.Status.MaterialInterlock"
   SymbolicIOField "valOutput2MaterialSupply2Low" at 280,150 size 220x25; TextOn '1'; TextOff '0'; TextList "MaterialInterlock_LabelSupply_NotLow"
      ProcessValue <- "PackTags.Status.MaterialInterlock"
   TextField "fraEquipmentInterlock" at 555,15 size 535x173; Text 'Equipment Interlock'
   TextField "txtEquipmentInterlockStarved" at 565,55 size 220x25; Text 'Upstream starved: / Zuführung leer: / Upstream Starved ..........'
   TextField "txtEquipmentInterlockBlocked" at 565,85 size 220x25; Text 'Downstream blocked: / Ausgabe blockiert:'
   GraphicIOField "valOutputtxtEquipmentInterlockStarved" at 790,55 size 25x25; PictureOff "PilotLight_Square_GN_Off_256c"; PictureOn "PilotLight_Square_R_On_256c"
      ProcessValue <- "PackTags.Status.EquipmentInterlock.Starved"
   GraphicIOField "valOutputtxtEquipmentInterlockBlocked" at 790,85 size 25x25; PictureOff "PilotLight_Square_GN_Off_256c"; PictureOn "PilotLight_Square_R_On_256c"
      ProcessValue <- "PackTags.Status.EquipmentInterlock.Blocked"

screen "1081_OMACStateModel" 1280x715, template "1xxx_MachineControl"
   ScreenModuleView "fcpOmacStateModel" at 5,5 size 1100x550; ScreenModuleType ""
      Guid_{11997190-30448} <- "PackTags.Admin.StatesDisabled"
      Guid_{11997190-30489} <- "PackTags.Status.StateCurrent"
   Rectangle "recBaseScreenLocked" at 0,0 size 1280x708
      Visibility <- "bo_System_BaseScreenLocked"

